   MV_MV22_CV1 : PlantItem := (CW := 2#0000_0000_0000_0000_0000_0000_1000_0001, DriveBits := 1);   // MV22_CV1
   MV_MV22_CV1_RawOutput : ALIAS FOR Remote_IO:12:O.Data.11;   // MV_MV22_CV1 MV22 coolant SOV
   MV_MV22_Filling_Pulse : BOOL;
   MV_MV22_Filling_PulseLevel : DINT := 252;
   MV_MV22_LTX07_AI : PlantItem := (CW := 2#0000_0000_0000_0000_1000_0000_0000_0000, CheckTime := 10, CheckTimer := 10, Scaled := 5.5534997, RawInput := 7064.0);   // MV22_LTX07
   MV_MV22_LTX07_AI_RawInput : ALIAS FOR Remote_IO:10:I.Ch05Data;   // Real Analog Input , Do Not Use In Code
   MV_MV22_LTX07_TrueLevel : REAL := 251.42085;
   MV_MV22_LTX07_TruePressure : REAL := 5.5534997;
   MV_MV22_Open_Vent_ALRM : ALARM_DIGITAL;
   MV_MV22_ProxiesOK : BOOL;
   MV_MV22_PTX01_AI : PlantItem := (CW := 2#0000_0000_0000_0000_1000_0000_0000_0000, CheckTime := 10, CheckTimer := 10, Scaled := -0.060749996, RawInput := 3946.0);   // MV22_PTX01
   MV_MV22_PTX01_AI_RawInput : ALIAS FOR Remote_IO:10:I.Ch02Data;   // Real Analog Input , Do Not Use In Code
   MV_MV22_PurgeAfterCIP : BOOL;
   MV_MV22_RTD1_AI : PlantItem := (CW := 2#0000_0000_0000_0000_1000_0000_0000_0000, CheckTime := 10, CheckTimer := 10, Scaled := -0.19999886, RawInput := -2.0);   // MV22_RTD1
   MV_MV22_RTD1_AI_RawInput : ALIAS FOR Remote_IO:5:I.Ch3Data;   // Real Analog Input , Do Not Use In Code
   MV_MV22_TP_CaskDepressure : BOOL;
   MV_MV22_TP_CaskEmptying : BOOL;
   MV_MV22_TP_CaskFilling : BOOL;
   MV_MV22_TP_CaskPreEmptyPressure : BOOL;
   MV_MV22_TP_CaskPrePressure : BOOL;
   MV_MV22_TP_CaskPressureDelay : BOOL;
   MV_MV22_TP_CaskPurgeFromTop : BOOL;
   MV_MV22_TP_CaskReadyToFill : BOOL;
   MV_MV22_TP_CaskStorage : BOOL;
   MV_MV22_TP_CO2_Debounce_Timer : TIMER := (PRE := 5000);
   MV_MV22_TP_CO2_Debounce_Timer_1 : TIMER := (PRE := 5000);
   MV_MV22_TP_CO2_HSL_Pressure : REAL := 16.0;
   MV_MV22_TP_CO2_HSL_Storage : REAL := 10.5;
   MV_MV22_TP_CO2_HSL_Timer : TIMER := (PRE := 5000, ACC := 5000, EN := 1, DN := 1);
   MV_MV22_TP_CO2_LSL_pressure : DINT := 9;
   MV_MV22_TP_CO2_LSL_pressure_1 : REAL := 2.0;
   MV_MV22_TP_CO2_LSL_storage : REAL := 9.5;
   MV_MV22_TP_CO2_LSL_Timer : TIMER := (PRE := 5000);
   MV_MV22_TP_CO2_Overshoot_pressure : DINT := 4;
   MV_MV22_TP_CO2_Pulse_Debounce_Timer : TIMER := (PRE := 5000);
   MV_MV22_TP_Command : DINT;
   MV_MV22_TP_DAL_Chase_Cask : BOOL;
   MV_MV22_TP_DAL_Chase_KB : BOOL;
   MV_MV22_TP_DAL_Chase_Time : TIMER := (PRE := 90000);
   MV_MV22_TP_Dirty : BOOL;
   MV_MV22_TP_DrainDown : BOOL;
   MV_MV22_TP_Emptying_Level_Setpoint : REAL := -260.0;
   MV_MV22_TP_Error_String : STRING;
   MV_MV22_TP_Faulted : BOOL;
   MV_MV22_TP_Fill_Pulse_OFF_Timer : TIMER := (PRE := 15000);
   MV_MV22_TP_Fill_Pulse_ON_Timer : TIMER := (PRE := 30000);
   MV_MV22_TP_Held : BOOL;
   MV_MV22_TP_Idle : BOOL;
   MV_MV22_TP_Initial_DAL_Chase_Cask : BOOL;
   MV_MV22_TP_Initial_DAL_Chase_KB : BOOL;
   MV_MV22_TP_KBDepressure : BOOL;
   MV_MV22_TP_KBEmptying : BOOL;
   MV_MV22_TP_KBFilling : BOOL;
   MV_MV22_TP_KBFilling_M : BOOL;
   MV_MV22_TP_KBFillingBuildPressure : BOOL;
   MV_MV22_TP_KBPreEmptyPressure : BOOL;
   MV_MV22_TP_KBPrePressurise : BOOL;
   MV_MV22_TP_KBPurgeFromTop : BOOL;
   MV_MV22_TP_KBPurgeTimer : TIMER;
   MV_MV22_TP_KBStorage : BOOL := 1;
   MV_MV22_TP_LowerLimit : REAL := 8.0;
   MV_MV22_TP_NotIdle : BOOL := 1;
   MV_MV22_TP_ONS : BOOL;
   MV_MV22_TP_ONS_1 : BOOL;
   MV_MV22_TP_PrePressure : BOOL;
   MV_MV22_TP_Prompt : DINT := 2;
   MV_MV22_TP_Proxy_Delay_Made : TIMER := (PRE := 2000);
   MV_MV22_TP_Proxy_Delay_NOT_MADE : TIMER := (PRE := 2000, ACC := 2000, EN := 1, DN := 1);
   MV_MV22_TP_Pulse : BOOL;
   MV_MV22_TP_ReadyToFillKB : BOOL;
   MV_MV22_TP_ReadyToFillKB_M : BOOL;
   MV_MV22_TP_Running : BOOL := 1;
   MV_MV22_TP_SeatClean_Delay : TIMER;
   MV_MV22_TP_SeatClean_Pulse : TIMER;
   MV_MV22_TP_Setpoint : REAL := 10.0;
   MV_MV22_TP_Status : DINT := 1;   // 0 = Idle, 1 = Running, 2 = Held, 3 = Faulted
   MV_MV22_TP_Step : DINT := 50;
   MV_MV22_TP_Steptime : DINT := 3562924;
   MV_MV22_TP_Steptime_String : STRING := '989:42:06';
   MV_MV22_TP_Steptime_String_1 : STRING;
   MV_MV22_TP_SteptimeRunning : DINT := 11;
   MV_MV22_TP_TimeLeft : DINT;
   MV_MV22_TP_TimeLeft_msec : DINT := 1;
   MV_MV22_TP_TimeLeftStr : STRING;
   MV_MV22_TP_UpperLimit : REAL := 12.0;
   MV_MV22_TP_Vent : BOOL;
   MV_MV22_TP_VentPressure : REAL;
   MV_MV22_TPLastStep : DINT := 50;
   MV_MV22_Transfer_StartLevel : REAL;
   MV_MV22_Transferred_Level : REAL := 95.31006;
   MV_MV22R : PlantItem := (CW := 2#0000_0000_0000_0010_0000_1100_0100_0001, CheckTime := 8, DriveBits := 1);   // MV22R
   MV_MV22R_ALARM : ALARM_DIGITAL;
   MV_MV22R_D : ALIAS FOR Remote_IO:14:O.Data.11;   // Rouser drive MV22
   MV_MV22R_R : ALIAS FOR Remote_IO:15:I.Data.27;   // MV22 Rouser running signal
   MV_MV23_CV1 : PlantItem;   // MV23_CV1
   MV_MV23_CV1_RawOutput : ALIAS FOR Remote_IO:12:O.Data.12;   // MV_MV23_CV1 MV23 coolant SOV
   MV_MV23_RTD1_AI : PlantItem := (CW := 2#0000_0000_0000_0000_1000_0000_0000_0000, CheckTime := 10, CheckTimer := 10, Scaled := 8.300001, RawInput := 83.0);   // MV23_RTD1
   MV_MV23_RTD1_AI_RawInput : ALIAS FOR Remote_IO:5:I.Ch4Data;   // Real Analog Input , Do Not Use In Code
   MV_MV23R : PlantItem := (CW := 2#0000_0000_0000_0010_0000_1100_0000_0000, CheckTime := 8, CheckTimer := 8);   // MV23R
   MV_MV23R_ALARM : ALARM_DIGITAL;
   MV_MV23R_D : ALIAS FOR Remote_IO:14:O.Data.12;   // Rouser drive MV23
   MV_MV23R_R : ALIAS FOR Remote_IO:15:I.Data.28;   // MV23 Rouser running signal
   MV_MV2_CV1 : PlantItem;   // MV2_CV1
   MV_MV2_CV1_RawOutput : ALIAS FOR Remote_IO:11:O.Data.1;   // MV_MV2_CV1
   MV_MV2_RTD1_AI : PlantItem := (CW := 2#0000_0000_0000_0000_1000_0000_0000_0000, CheckTime := 10, CheckTimer := 10, Scaled := 8.200001, RawInput := 82.0);   // MV2_RTD1
   MV_MV2_RTD1_AI_RawInput : ALIAS FOR Remote_IO:1:I.Ch1Data;   // Real Analog Input , Do Not Use In Code
   MV_MV2R : PlantItem := (CW := 2#0000_0000_0000_0011_0000_1100_0000_0000, CheckTime := 8, CheckTimer := 8);   // MV2R
   MV_MV2R_ALARM : ALARM_DIGITAL;
   MV_MV2R_ALM : ALARM_DIGITAL;
   MV_MV2R_D : ALIAS FOR Remote_IO:13:O.Data.1;
   MV_MV2R_R : ALIAS FOR Remote_IO:15:I.Data.1;   // MV2 Rouser running signal
   MV_MV30_CV1 : PlantItem;   // MV30_CV1
   MV_MV30_CV1_RawOutput : ALIAS FOR Remote_IO:12:O.Data.3;   // MV_MV30_CV1 MV30 coolant SOV
   MV_MV30_RTD1_AI : PlantItem := (CW := 2#0000_0000_0000_0000_1000_0000_0000_0000, CheckTime := 10, CheckTimer := 10, Scaled := 21.900002, RawInput := 219.0);   // MV30_RTD1
   MV_MV30_RTD1_AI_RawInput : ALIAS FOR Remote_IO:4:I.Ch1Data;   // Real Analog Input , Do Not Use In Code
   MV_MV30R : PlantItem := (CW := 2#0000_0000_0000_0010_0000_1100_0000_0000, CheckTime := 8, CheckTimer := 8);   // MV30R
   MV_MV30R_ALARM : ALARM_DIGITAL;
   MV_MV30R_D : ALIAS FOR Remote_IO:14:O.Data.3;   // Rouser drive MV30
   MV_MV30R_R : ALIAS FOR Remote_IO:15:I.Data.19;   // MV30 Rouser running signal
   MV_MV31_CV1 : PlantItem;   // MV31_CV1
   MV_MV31_CV1_RawOutput : ALIAS FOR Remote_IO:12:O.Data.4;   // MV_MV31_CV1 MV31coolant SOV
   MV_MV31_RTD1_AI : PlantItem := (CW := 2#0000_0000_0000_0000_1000_0000_0000_0000, CheckTime := 10, CheckTimer := 10, Scaled := 6.300001, RawInput := 63.0);   // MV31_RTD1
   MV_MV31_RTD1_AI_RawInput : ALIAS FOR Remote_IO:4:I.Ch2Data;   // Real Analog Input , Do Not Use In Code
   MV_MV31R : PlantItem := (CW := 2#0000_0000_0000_0010_0000_1100_0000_0000, CheckTime := 8, CheckTimer := 8);   // MV31R
   MV_MV31R_ALARM : ALARM_DIGITAL;
   MV_MV31R_D : ALIAS FOR Remote_IO:14:O.Data.4;   // Rouser drive MV31
   MV_MV31R_R : ALIAS FOR Remote_IO:15:I.Data.20;   // MV31 Rouser running signal
   MV_MV32_CV1 : PlantItem;   // MV32_CV1
   MV_MV32_CV1_RawOutput : ALIAS FOR Remote_IO:12:O.Data.5;   // MV_MV32_CV1 MV32 coolant SOV
   MV_MV32_RTD1_AI : PlantItem := (CW := 2#0000_0000_0000_0000_1000_0000_0000_0000, CheckTime := 10, CheckTimer := 10, Scaled := 22.0, RawInput := 220.0);   // MV32_RTD1
   MV_MV32_RTD1_AI_RawInput : ALIAS FOR Remote_IO:4:I.Ch3Data;   // Real Analog Input , Do Not Use In Code
   MV_MV32R : PlantItem := (CW := 2#0000_0000_0000_0010_0000_1100_0000_0000, CheckTime := 8, CheckTimer := 8);   // MV32R
   MV_MV32R_ALARM : ALARM_DIGITAL;
   MV_MV32R_D : ALIAS FOR Remote_IO:14:O.Data.5;   // Rouser drive MV32
   MV_MV32R_R : ALIAS FOR Remote_IO:15:I.Data.21;   // MV32 Rouser running signal
   MV_MV33_CV1 : PlantItem;   // MV33_CV1
   MV_MV33_CV1_RawOutput : ALIAS FOR Remote_IO:12:O.Data.6;   // MV_MV33_CV1 MV33 coolant SOV
   MV_MV33_RTD1_AI : PlantItem := (CW := 2#0000_0000_0000_0000_1000_0000_0000_0000, CheckTime := 10, CheckTimer := 10, Scaled := 8.1, RawInput := 81.0);   // MV33_RTD1
   MV_MV33_RTD1_AI_RawInput : ALIAS FOR Remote_IO:4:I.Ch4Data;   // Real Analog Input , Do Not Use In Code
   MV_MV33R : PlantItem := (CW := 2#0000_0000_0000_0010_0000_1100_0000_0000, CheckTime := 8, CheckTimer := 8);   // MV33R
   MV_MV33R_ALARM : ALARM_DIGITAL;
   MV_MV33R_D : ALIAS FOR Remote_IO:14:O.Data.6;   // Rouser drive MV33
   MV_MV33R_R : ALIAS FOR Remote_IO:15:I.Data.22;   // MV33 Rouser running signal
   MV_MV34_CV1 : PlantItem;   // MV34_CV1
   MV_MV34_CV1_RawOutput : ALIAS FOR Remote_IO:12:O.Data.7;   // MV_MV34_CV1 MV34 coolant SOV
   MV_MV34_RTD1_AI : PlantItem := (CW := 2#0000_0000_0000_0000_1000_0000_0000_0000, CheckTime := 10, CheckTimer := 10, Scaled := 22.100002, RawInput := 221.0);   // MV34_RTD1
   MV_MV34_RTD1_AI_RawInput : ALIAS FOR Remote_IO:4:I.Ch5Data;   // Real Analog Input , Do Not Use In Code
   MV_MV34R : PlantItem := (CW := 2#0000_0000_0000_0010_0000_1100_0000_0000, CheckTime := 8, CheckTimer := 8);   // MV34R
   MV_MV34R_ALARM : ALARM_DIGITAL;
   MV_MV34R_D : ALIAS FOR Remote_IO:14:O.Data.7;   // Rouser drive MV34
   MV_MV34R_R : ALIAS FOR Remote_IO:15:I.Data.23;   // MV34 Rouser running signal
   MV_MV35_CV1 : PlantItem;   // MV35_CV1
   MV_MV35_CV1_RawOutput : ALIAS FOR Remote_IO:12:O.Data.8;   // MV_MV35_CV1 MV35 coolant SOV
   MV_MV35_RTD1_AI : PlantItem := (CW := 2#0000_0000_0000_0000_1000_0000_0000_0000, CheckTime := 10, CheckTimer := 10, Scaled := 22.8, RawInput := 228.0);   // MV35_RTD1
   MV_MV35_RTD1_AI_RawInput : ALIAS FOR Remote_IO:5:I.Ch0Data;   // Real Analog Input , Do Not Use In Code
   MV_MV35R : PlantItem := (CW := 2#0000_0000_0000_0010_0000_1100_0000_0000, CheckTime := 8, CheckTimer := 8);   // MV35R
   MV_MV35R_ALARM : ALARM_DIGITAL;
   MV_MV35R_D : ALIAS FOR Remote_IO:14:O.Data.8;   // Rouser drive MV35
   MV_MV35R_R : ALIAS FOR Remote_IO:15:I.Data.24;   // MV35 Rouser running signal
   MV_MV36_AV01 : PlantItem;   // MV36_AV01
   MV_MV36_AV01_RawOutput : ALIAS FOR Remote_IO:16:O.Data.0;   // MV_MV36_AV01
   MV_MV36_TTX01_AI : PlantItem := (CW := 2#0000_0000_0000_0000_1000_0000_0000_0000, CheckTime := 10, CheckTimer := 10, Scaled := 8.096876, RawInput := 9791.0);   // MV36_TTX01
   MV_MV36_TTX01_AI_RawInput : ALIAS FOR Remote_IO:7:I.Ch00Data;   // Real Analog Input , Do Not Use In Code
   MV_MV37_AV01 : PlantItem := (CW := 2#0000_0000_0000_0000_0000_0000_0010_0000);   // MV37_AV01
   MV_MV37_AV01_RawOutput : ALIAS FOR Remote_IO:16:O.Data.1;   // MV_MV37_AV01 MV37 coolant SOV
   MV_MV37_TTX01_AI : PlantItem := (CW := 2#0000_0000_0000_0000_1000_0000_0000_0000, CheckTime := 10, CheckTimer := 10, Scaled := -1.4093752, RawInput := 6749.0);   // MV37_TTX01
   MV_MV37_TTX01_AI_RawInput : ALIAS FOR Remote_IO:7:I.Ch01Data;   // Real Analog Input , Do Not Use In Code
   MV_MV38_AV01 : PlantItem;   // MV38_AV01
   MV_MV38_AV01_RawOutput : ALIAS FOR Remote_IO:16:O.Data.2;   // MV_MV38_AV01 MV38 coolant SOV
   MV_MV38_TTX01_AI : PlantItem := (CW := 2#0000_0000_0000_0000_1000_0000_0000_0000, CheckTime := 10, CheckTimer := 10, Scaled := 8.1, RawInput := 9792.0);   // MV38_TTX01
   MV_MV38_TTX01_AI_RawInput : ALIAS FOR Remote_IO:7:I.Ch02Data;   // Real Analog Input , Do Not Use In Code
   MV_MV39_AV01 : PlantItem;   // MV39_AV01
   MV_MV39_AV01_RawOutput : ALIAS FOR Remote_IO:16:O.Data.3;   // MV_MV39_AV01 MV39 coolant SOV
   MV_MV39_TTX01_AI : PlantItem := (CW := 2#0000_0000_0000_0000_1000_0000_0000_0000, CheckTime := 10, CheckTimer := 10, Scaled := -1.4437494, RawInput := 6738.0);   // MV39_TTX01
   MV_MV39_TTX01_AI_RawInput : ALIAS FOR Remote_IO:7:I.Ch03Data;   // Real Analog Input , Do Not Use In Code
   MV_MV3_CV1 : PlantItem;   // MV3_CV1
   MV_MV3_CV1_RawOutput : ALIAS FOR Remote_IO:11:O.Data.2;   // MV_MV3_CV1 MV3 coolant SOV
   MV_MV3_RTD1_AI : PlantItem := (CW := 2#0000_0000_0000_0000_1000_0000_0000_0000, CheckTime := 10, CheckTimer := 10, Scaled := 8.1, RawInput := 81.0);   // MV3_RTD1
   MV_MV3_RTD1_AI_RawInput : ALIAS FOR Remote_IO:1:I.Ch2Data;   // Real Analog Input , Do Not Use In Code
   MV_MV3R : PlantItem := (CW := 2#0000_0000_0000_0010_0000_1100_0000_0000, CheckTime := 8, CheckTimer := 8);   // MV3R
   MV_MV3R_ALARM : ALARM_DIGITAL;
   MV_MV3R_D : ALIAS FOR Remote_IO:13:O.Data.2;   // Rouser drive MV3
   MV_MV3R_R : ALIAS FOR Remote_IO:15:I.Data.2;   // MV3 Rouser running signal
   MV_MV40_AV01 : PlantItem;   // MV40_AV01
   MV_MV40_AV01_RawOutput : ALIAS FOR Remote_IO:16:O.Data.4;   // MV_MV40_AV01 MV40 coolant SOV
   MV_MV40_TTX01_AI : PlantItem := (CW := 2#0000_0000_0000_0000_1000_0000_0000_0000, CheckTime := 10, CheckTimer := 10, Scaled := 7.7562504, RawInput := 9682.0);   // MV40_TTX01
   MV_MV40_TTX01_AI_RawInput : ALIAS FOR Remote_IO:7:I.Ch04Data;   // Real Analog Input , Do Not Use In Code
   MV_MV41_AV01 : PlantItem;   // MV41_AV01
   MV_MV41_AV01_RawOutput : ALIAS FOR Remote_IO:16:O.Data.5;   // MV_MV41_AV01 MV41 coolant SOV
   MV_MV41_TTX01_AI : PlantItem := (CW := 2#0000_0000_0000_0000_1000_0000_0000_0000, CheckTime := 10, CheckTimer := 10, Scaled := 7.846876, RawInput := 9711.0);   // MV41_TTX01
   MV_MV41_TTX01_AI_RawInput : ALIAS FOR Remote_IO:7:I.Ch05Data;   // Real Analog Input , Do Not Use In Code
   MV_MV42_AV01 : PlantItem;   // MV42_AV01
   MV_MV42_AV01_RawOutput : ALIAS FOR Remote_IO:16:O.Data.6;   // MV_MV42_AV01 MV42 coolant SOV
   MV_MV42_TTX01_AI : PlantItem := (CW := 2#0000_0000_0000_0000_1000_0000_0000_0000, CheckTime := 10, CheckTimer := 10, Scaled := 21.015625, RawInput := 13925.0);   // MV42_TTX01
   MV_MV42_TTX01_AI_RawInput : ALIAS FOR Remote_IO:7:I.Ch06Data;   // Real Analog Input , Do Not Use In Code
   MV_MV43_AV01 : PlantItem;   // MV43_AV01
   MV_MV43_AV01_RawOutput : ALIAS FOR Remote_IO:16:O.Data.7;   // MV_MV43_AV01 MV43 coolant SOV
   MV_MV43_TTX01_AI : PlantItem := (CW := 2#0000_0000_0000_0000_1000_0000_0000_0000, CheckTime := 10, CheckTimer := 10, Scaled := 21.221876, RawInput := 13991.0);   // MV43_TTX01
   MV_MV43_TTX01_AI_RawInput : ALIAS FOR Remote_IO:7:I.Ch07Data;   // Real Analog Input , Do Not Use In Code
   MV_MV44_AV01 : PlantItem;   // MV44_AV01
   MV_MV44_AV01_RawOutput : ALIAS FOR Remote_IO:16:O.Data.8;   // MV_MV44_AV01 MV44 coolant SOV
   MV_MV44_TTX01_AI : PlantItem := (CW := 2#0000_0000_0000_0000_1000_0000_0000_0000, CheckTime := 10, CheckTimer := 10, Scaled := 21.075, RawInput := 13944.0);   // MV44_TTX01
   MV_MV44_TTX01_AI_RawInput : ALIAS FOR Remote_IO:7:I.Ch08Data;   // Real Analog Input , Do Not Use In Code
   MV_MV45_AV01 : PlantItem;   // MV45_AV01
   MV_MV45_AV01_RawOutput : ALIAS FOR Remote_IO:16:O.Data.9;   // MV_MV45_AV01 MV45 coolant SOV
   MV_MV45_TTX01_AI : PlantItem := (CW := 2#0000_0000_0000_0000_1000_0000_0000_0000, CheckTime := 10, CheckTimer := 10, Scaled := 7.778126, RawInput := 9689.0);   // MV45_TTX01
   MV_MV45_TTX01_AI_RawInput : ALIAS FOR Remote_IO:7:I.Ch09Data;   // Real Analog Input , Do Not Use In Code
   MV_MV46_AV01 : PlantItem;   // MV46_AV01
   MV_MV46_AV01_RawOutput : ALIAS FOR Remote_IO:16:O.Data.10;   // MV_MV46_AV01 MV46 coolant SOV
   MV_MV46_TTX01_AI : PlantItem := (CW := 2#0000_0000_0000_0000_1000_0000_0000_0000, CheckTime := 10, CheckTimer := 10, Scaled := 21.25625, RawInput := 14002.0);   // MV46_TTX01
   MV_MV46_TTX01_AI_RawInput : ALIAS FOR Remote_IO:7:I.Ch10Data;   // Real Analog Input , Do Not Use In Code
   MV_MV47_AV01 : PlantItem := (CW := 2#0000_0000_0000_0000_0000_0000_1000_0001, DriveBits := 1);   // MV47_AV01
   MV_MV47_AV01_RawOutput : ALIAS FOR Remote_IO:16:O.Data.11;   // MV_MV47_AV01 MV47 coolant SOV
   MV_MV47_TTX01_AI : PlantItem := (CW := 2#0000_0000_0000_0000_1000_0000_0000_0000, CheckTime := 10, CheckTimer := 10, Scaled := -1.2468748, RawInput := 6801.0);   // MV47_TTX01
   MV_MV47_TTX01_AI_RawInput : ALIAS FOR Remote_IO:7:I.Ch11Data;   // Real Analog Input , Do Not Use In Code
   MV_MV4_CV1 : PlantItem;   // MV4_CV1
   MV_MV4_CV1_RawOutput : ALIAS FOR Remote_IO:11:O.Data.3;   // MV_MV4_CV1 MV4 coolant SOV
   MV_MV4_RTD1_AI : PlantItem := (CW := 2#0000_0000_0000_0000_1000_0000_0000_0000, CheckTime := 10, CheckTimer := 10, Scaled := 8.0, RawInput := 80.0);   // MV4_RTD1
   MV_MV4_RTD1_AI_RawInput : ALIAS FOR Remote_IO:1:I.Ch3Data;   // Real Analog Input , Do Not Use In Code
   MV_MV4R : PlantItem := (CW := 2#0000_0000_0000_0010_0000_1100_0000_0000, CheckTime := 8, CheckTimer := 8);   // MV4R
   MV_MV4R_ALARM : ALARM_DIGITAL;
   MV_MV4R_D : ALIAS FOR Remote_IO:13:O.Data.3;   // Rouser drive MV4
   MV_MV4R_R : ALIAS FOR Remote_IO:15:I.Data.3;   // MV4 Rouser running signal
   MV_MV5_CV1 : PlantItem;   // MV5_CV1
   MV_MV5_CV1_RawOutput : ALIAS FOR Remote_IO:11:O.Data.4;   // MV_MV5_CV1 MV5 coolant SOV
   MV_MV5_RTD1_AI : PlantItem := (CW := 2#0000_0000_0000_0000_1000_0000_0000_0000, CheckTime := 10, CheckTimer := 10, Scaled := 8.200001, RawInput := 82.0);   // MV5_RTD1
   MV_MV5_RTD1_AI_RawInput : ALIAS FOR Remote_IO:1:I.Ch4Data;   // Real Analog Input , Do Not Use In Code
   MV_MV5R : PlantItem := (CW := 2#0000_0000_0000_0010_0000_1100_0000_0000, CheckTime := 8, CheckTimer := 8);   // MV5R
   MV_MV5R_ALARM : ALARM_DIGITAL;
   MV_MV5R_D : ALIAS FOR Remote_IO:13:O.Data.4;   // Rouser drive MV5
   MV_MV5R_R : ALIAS FOR Remote_IO:15:I.Data.4;   // MV5 Rouser running signal
   MV_MV6_CV1 : PlantItem;   // MV6_CV1
   MV_MV6_CV1_RawOutput : ALIAS FOR Remote_IO:11:O.Data.5;   // MV_MV6_CV1 MV6 coolant SOV
   MV_MV6_RTD1_AI : PlantItem := (CW := 2#0000_0000_0000_0000_1000_0000_0000_0000, CheckTime := 10, CheckTimer := 10, Scaled := 25.100002, RawInput := 251.0);   // MV6_RTD1
   MV_MV6_RTD1_AI_RawInput : ALIAS FOR Remote_IO:1:I.Ch5Data;   // Real Analog Input , Do Not Use In Code
   MV_MV6R : PlantItem := (CW := 2#0000_0000_0000_0010_0000_1100_0000_0000, CheckTime := 8, CheckTimer := 8);   // MV6R
   MV_MV6R_ALARM : ALARM_DIGITAL;
   MV_MV6R_D : ALIAS FOR Remote_IO:13:O.Data.5;   // Rouser drive MV6
   MV_MV6R_R : ALIAS FOR Remote_IO:15:I.Data.5;   // MV6 Rouser running signal
   MV_MV7_CV1 : PlantItem;   // MV7_CV1
   MV_MV7_CV1_RawOutput : ALIAS FOR Remote_IO:11:O.Data.6;   // MV_MV7_CV1 MV7 coolant SOV
   MV_MV7_RTD1_AI : PlantItem := (CW := 2#0000_0000_0000_0000_1000_0000_0000_0000, CheckTime := 10, CheckTimer := 10, Scaled := 8.200001, RawInput := 82.0);   // MV7_RTD1
   MV_MV7_RTD1_AI_RawInput : ALIAS FOR Remote_IO:2:I.Ch0Data;   // Real Analog Input , Do Not Use In Code
   MV_MV7R : PlantItem := (CW := 2#0000_0000_0000_0010_0000_1100_0000_0000, CheckTime := 8, CheckTimer := 8);   // MV7R
   MV_MV7R_ALARM : ALARM_DIGITAL;
   MV_MV7R_D : ALIAS FOR Remote_IO:13:O.Data.6;   // Rouser drive MV7
   MV_MV7R_R : ALIAS FOR Remote_IO:15:I.Data.6;   // MV7 Rouser running signal
   MV_MV8_CV1 : PlantItem := (CW := 2#0000_0000_0000_0000_0000_0000_1000_0001, DriveBits := 1);   // MV8_CV1
   MV_MV8_CV1_RawOutput : ALIAS FOR Remote_IO:11:O.Data.7;   // MV_MV8_CV1 MV8 coolant SOV
   MV_MV8_RTD1_AI : PlantItem := (CW := 2#0000_0000_0000_0000_1000_0000_0000_0000, CheckTime := 10, CheckTimer := 10, Scaled := 9.700001, RawInput := 97.0);   // MV8_RTD1
   MV_MV8_RTD1_AI_RawInput : ALIAS FOR Remote_IO:2:I.Ch1Data;   // Real Analog Input , Do Not Use In Code
   MV_MV8R : PlantItem := (CW := 2#0000_0000_0000_0010_0000_1100_0000_0000, CheckTime := 8, CheckTimer := 8);   // MV8R
   MV_MV8R_ALARM : ALARM_DIGITAL;
   MV_MV8R_D : ALIAS FOR Remote_IO:13:O.Data.7;   // Rouser drive MV8
   MV_MV8R_R : ALIAS FOR Remote_IO:15:I.Data.7;   // MV8 Rouser running signal
   MV_MV9_CV1 : PlantItem := (CW := 2#0000_0000_0000_0000_0000_0000_0010_0000);   // MV9_CV1
   MV_MV9_CV1_RawOutput : ALIAS FOR Remote_IO:11:O.Data.8;   // MV_MV9_CV1 MV9 coolant SOV
   MV_MV9_RTD1_AI : PlantItem := (CW := 2#0000_0000_0000_0000_1000_0000_0000_0000, CheckTime := 10, CheckTimer := 10, Scaled := 26.400002, RawInput := 264.0);   // MV9_RTD1
   MV_MV9_RTD1_AI_RawInput : ALIAS FOR Remote_IO:2:I.Ch2Data;   // Real Analog Input , Do Not Use In Code
   MV_MV9R : PlantItem := (CW := 2#0000_0000_0000_0010_0000_1100_0000_0000, CheckTime := 8, CheckTimer := 8);   // MV9R
   MV_MV9R_ALARM : ALARM_DIGITAL;
   MV_MV9R_D : ALIAS FOR Remote_IO:13:O.Data.8;   // Rouser drive MV9
   MV_MV9R_R : ALIAS FOR Remote_IO:15:I.Data.8;   // MV9 Rouser running signal
   MV_N101 : INT[255] := ([0] := 152, [1] := -15, [2] := -15, [3] := 1680, [4] := 5280, [5] := 2950, [6] := 463, [7] := 124, [8] := 7, [9] := 3, [10] := 110, [11] := -13);   // AT INT Fermentation control integer workspace
        [1]   // Setpoint at previous breakpoint
        [4]   // Next breakpoint time
        [6]   // Temporary result register
        [5]   // Time since last B.P in 1/10 hour
        [3]   // Previous breakpoint time
        [0]   // Attemporation Control Loop Current Vessel File Pointer
        [7]   // Pointer to vessel's data file
        [8]   // Number of open cooling valves
        [11]   // Temp.register
        [2]   // Setpoint at next breakpoint
        [9]   // Rouser operation temperature
   MV_N104 : INT[255] := ([0] := -32768, [1] := -32768, [2] := -32768, [3] := -32768, [4] := -32768, [5] := -32768, [6] := -32768, [7] := -32768, [8] := -32768, [9] := -32768, [10] := -32768, [11] := -32768, [12] := -32768, [13] := -32768, [14] := -32768, [15] := -32768, [16] := -32768, [17] := -32768, [18] := -32768, [19] := -32768, [20] := -32768, [21] := -32768, [22] := -32768, [23] := -32768, [24] := -32768);   // MV_PC_BUF PC>PLC Attemporation Control Command Buf fer File
        [10]   // PC>PLC FV System Command Buffer Breakpoint E Temperature Setpoint
        [12]   // PC>PLC FV System Command Buffer Breakpoint F Temperature Setpoint
        [14]   // PC>PLC FV System Command Buffer Breakpoint G Temperature Setpoint
        [1]   // PC>PLC Attemporation System Command Buffer Breakpoint A Time
        [15]   // PC>PLC FV System Command Buffer Profile Control / Configuration Flags
        [15].6   // FV System PC Command Buffer Control Flags 1=Wait for yeast required
        [2]   // PC>PLC FV System Command Buffer Breakpoint A Temperature Setpoint
        [4]   // PC>PLC FV System Command Buffer Breakpoint B Temperature Setpoint
        [6]   // PC>PLC FV System Command Buffer Breakpoint C Temperature Setpoint
        [15].4   // FV System PC Command Buffer Control Flags 1=Ageing Profile
        [8]   // PC>PLC FV System Command Buffer Breakpoint D Temperature Setpoint
        [23]   // PC>PLC AT System Command Buffer Command Type 1=Start,2=Stop 3=Modify Control
        [0]   // PC>PLC Attempotation System Vessel Number 29-56,94 = MV1-MV23 336-347 = MV36-47
        [15].5   // FV System PC Command Buffer Control Flags 1=Conditioning Profile
        [11]   // PC>PLC FV System Command Buffer Breakpoint F Time
        [13]   // PC>PLC FV System Command Buffer Breakpoint G Time
        [24]   // Attemporation System PC Command Buffer Phase Number
        [16]   // PC>PLC FV System Command Buffer PC Private Flags
        [3]   // PC>PLC FV System Command Buffer Breakpoint B Time
        [5]   // PC>PLC FV System Command Buffer Breakpoint C Time
        [7]   // PC>PLC FV System Command Buffer Breakpoint D Time
        [9]   // PC>PLC FV System Command Buffer Breakpoint E Time
   MV_N105 : INT[255] := ([0] := 1025, [1] := 116, [3] := 45, [4] := 114);   // ROUSE_CTRL Rouser control progr am working regs
        [2]   // PC>PLC Rouser control Vessel number to be set to timed mode
        [0].0   // Rouser control 1 minute latch
        [0].10   // Rouser Control Hourly Latch
        [0].2   // Rouser Control Daily latch synchroniser
        [0].9   // Rouser Control Hourly latch synchroniser
        [4]   // Rouse control PC timed rouse request vessel pointer
        [1]   // Rouser control current vessel data file pointer
        [0].3   // Rouser Control Daily Latch
        [3]   // PC>PLC Rouser control Timed rouse duration
        [0].4   // Rouser control 1 minute latch synchroniser
   MV_N105_0_1_Output_Bit : BOOL;
   MV_N105_0_6_Output_Bit : BOOL;
   MV_N105_0_7_Output_Bit : BOOL;
   MV_N105_0_8_Output_Bit : BOOL;
   MV_N106 : INT[255] := ([0] := 33, [2] := 80, [3] := 1680, [4] := 80, [5] := 3360, [6] := 80, [7] := 5040, [8] := 80, [9] := 6720, [10] := 80, [11] := 8400, [12] := 80, [13] := 32767, [14] := 80, [15] := 148, [17] := -32767, [18] := -32767, [19] := 1680, [20] := 3171, [22] := 4639, [23] := 1, [24] := 10, [25] := 82, [26] := 80, [27] := 3171, [29] := 2, [30] := 24, [32] := 2, [34] := 2, [42] := 25640);   // ROUSE_BUFF Rouser control vesse l data buffer
        [24]   // Phase 0=off 8=Wait yeast 10=Maturation 11to16=Conditioning
        [32]   // Rouser control mode 0=Off 1=Continuous 2=Daily 3=Timed 4=Hourly
        [30].2   // Rouse required due to high temperature
        [29].1   // Current vessel deferred chilling enabled flag
        [30].0   // Current vessel cooling valve required to open
        [34]   // Saved rouser mode of operation
        [27]   // Current vessel elapsed time
        [15].7   // Profile control flag Rousing enabled
        [25]   // ACTUAL TEMPERATURE -DEGREES 'C'*10
        [30].1   // Rouser to run
        [31]   // Rouser run time remaining (minutes)
   MV_N110 : INT[255] := ([0] := 347, [2] := 100, [3] := 1200, [4] := 100, [5] := 1680, [6] := -15, [7] := 5280, [8] := -15, [9] := 7210, [10] := -15, [11] := 8340, [12] := -15, [13] := 32767, [14] := -15, [15] := 164, [17] := -32767, [18] := -32767, [19] := 1680, [20] := 1200, [21] := 2981, [22] := 6282, [23] := 1, [24] := 13, [25] := -13, [26] := -15, [27] := 4630, [29] := 257, [30] := 123, [32] := 2, [34] := 2, [40] := 2);   // MV DATA 0 CURRENT FV DATA
        [15].5   // Profile Control Flags : This is a Conditioning Profile
        [24]   // Phase 0=off 8=Wait yeast 9=Wait Fill 10=Maturation 11to16=Conditioning
        [15].9   // Current vessel deferred chilling manual override
        [22]   // Current FV total residence time
        [29].0   // PC TO SAVE TEMPERATURE DATA
        [40]   // Vessel RoutingStatus 0=Clean,1=Filling,2= Beer,3=Packng1,4=Pac kng2,5=Packng3,6=Ven ting,7=Dirty,8=CIP
        [15].4   // Profile Control Flags : This is a Maturation Profile
        [1]   // TEMPERATURE BREAKPOINT A. TIME 1/10 HOURS(ALWAYS=0)
        [11]   // TEMPERATURE BREAKPOINT F. TIME 1/10 HOURS(ALWAYS=0)
        [29].1   // Current vessel deferred chilling enabled flag
        [13]   // TEMPERATURE BREAKPOINT G. TIME 1/10 HOURS(ALWAYS=0)
        [3]   // TEMPERATURE BREAKPOINT B. TIME 1/10 HOURS(ALWAYS=0)
        [30].5   // Current vessel deferred chilling temp.high flag
        [30].3   // Current vessel deferred chilling active
        [5]   // TEMPERATURE BREAKPOINT C. TIME 1/10 HOURS(ALWAYS=0)
        [7]   // TEMPERATURE BREAKPOINT D. TIME 1/10 HOURS(ALWAYS=0)
        [9]   // TEMPERATURE BREAKPOINT E. TIME 1/10 HOURS(ALWAYS=0)
        [16].1   // Profile control flag Hold at B.P B
        [16].2   // Profile control flag Hold at B.P C
        [16].3   // Profile control flag Hold at B.P D
        [16].4   // Profile control flag Hold at B.P E
        [16].5   // Profile control flag Hold at B.P F
        [16].6   // Profile control flag Hold at B.P G
        [15].2   // PLC TO FOLLOW RAMP Breakpoints A to B
        [0]   // FV SYSTEM WORKING BUFFER VESSEL NUMBER
        [10]   // TEMPERATURE SETPOINT E. 1/10 DEGREE 'C'
        [12]   // TEMPERATURE SETPOINT F. 1/10 DEGREE 'C'
        [14]   // TEMPERATURE SETPOINT G. 1/10 DEGREE 'C'
        [21]   // Current vessel cold conditioning time
        [2]   // TEMPERATURE SETPOINT A. 1/10 DEGREE 'C'
        [30].4   // Current vessel final temp.reached
        [36]   // Current vessel time to deferred chlling start (hrs.x10)
        [4]   // TEMPERATURE SETPOINT B. 1/10 DEGREE 'C'
        [30].6   // Current vessel cold cond.temp.reached
        [6]   // TEMPERATURE SETPOINT C. 1/10 DEGREE 'C'
        [8]   // TEMPERATURE SETPOINT D. 1/10 DEGREE 'C'
        [15].3   // PLC TO USE CONE COOLING JACKET
        [25]   // ACTUAL TEMPERATURE -DEGREES 'C'*10
        [26]   // Calculated Setpoint 1/10 degrees C
        [44]   // Current vessel powder amount
        [20]   // Current FV warm conditioning time
        [29]   // FLAGS - PLC CONTROL
        [15]   // FLAGS-PROFILE CONTROL
        [28]   // CURRENT VOLUME HL*10
        [30].1   // Rouser required
        [27]   // CURRENT ELAPSED HOURS *10
        [30].0   // Cooling Valve to open
        [15].7   // PC>PLC Rousing enabled
        [43]   // Current vessel powder type
   MV_N111 : INT[50] := ([0] := 29, [2] := 80, [3] := 1200, [4] := 80, [5] := 1730, [6] := 80, [7] := 5040, [8] := 80, [9] := 6720, [10] := 80, [11] := 8400, [12] := 80, [13] := 32767, [14] := 80, [15] := 148, [17] := -32767, [18] := -32767, [19] := 1680, [20] := 311, [22] := 1947, [23] := 1, [24] := 10, [25] := 80, [26] := 80, [27] := 311, [30] := 19, [32] := 2, [34] := 2, [36] := 170, [42] := 25900);   // MV 1, CURRENT FV DATA
        [24]   // MV 1,Phase 0=off 8=Wait yeast 9=Wait Fill 10=Maturation 11to16=Conditioning
        [11]   // MV 1,TEMPERATURE BREAKPOINT F. TIME 1/10 HOURS(ALWAYS=0)
        [13]   // MV 1,TEMPERATURE BREAKPOINT G. TIME 1/10 HOURS(ALWAYS=0)
        [30].5   // MV 1,Current vessel deferred chilling temp.high flag
        [1]   // MV 1,TEMPERATURE BREAKPOINT A. TIME 1/10 HOURS(ALWAYS=0)
        [29].1   // MV 1,Current vessel deferred chilling enabled flag
        [3]   // MV 1,TEMPERATURE BREAKPOINT B. TIME 1/10 HOURS(ALWAYS=0)
        [5]   // MV 1,TEMPERATURE BREAKPOINT C. TIME 1/10 HOURS(ALWAYS=0)
        [36]   // MV 1,Current vessel time to deferred chlling start (hrs.x10)
        [15].5   // MV 1,Profile Control Flags : This is a Conditioning Profile
        [40]   // MV 1,Vessel RoutingStatus 0=Clean,1=Filling,2= Beer,3=Packng1,4=Pac kng2,5=Packng3,6=Ven ting,7=Dirty,8=CIP
        [15].7   // MV 1,PC>PLC Rousing enabled
        [43]   // MV 1,Current vessel powder type
        [15].4   // MV 1,Profile Control Flags : This is a Maturation Profile
        [16].1   // MV 1,Profile control flag Hold at B.P B
        [16].2   // MV 1,Profile control flag Hold at B.P C
        [10]   // MV 1,TEMPERATURE SETPOINT E. 1/10 DEGREE 'C'
        [7]   // MV 1,TEMPERATURE BREAKPOINT D. TIME 1/10 HOURS(ALWAYS=0)
        [12]   // MV 1,TEMPERATURE SETPOINT F. 1/10 DEGREE 'C'
        [14]   // MV 1,TEMPERATURE SETPOINT G. 1/10 DEGREE 'C'
        [9]   // MV 1,TEMPERATURE BREAKPOINT E. TIME 1/10 HOURS(ALWAYS=0)
        [0]   // MV 1,FV SYSTEM WORKING BUFFER VESSEL NUMBER
        [21]   // MV 1,Current vessel cold conditioning time
        [16].3   // MV 1,Profile control flag Hold at B.P D
        [2]   // MV 1,TEMPERATURE SETPOINT A. 1/10 DEGREE 'C'
        [30].3   // MV 1,Current vessel deferred chilling active
        [16].4   // MV 1,Profile control flag Hold at B.P E
        [30].4   // MV 1,Current vessel final temp.reached
        [16].5   // MV 1,Profile control flag Hold at B.P F
        [4]   // MV 1,TEMPERATURE SETPOINT B. 1/10 DEGREE 'C'
        [15].2   // MV 1,PLC TO FOLLOW RAMP Breakpoints A to B
        [20]   // MV 1,Current FV warm conditioning time
        [15].3   // MV 1,PLC TO USE CONE COOLING JACKET
        [15].9   // MV 1,Current vessel deferred chilling manual override
        [30].6   // MV 1,Current vessel cold cond.temp.reached
        [25]   // MV 1,ACTUAL TEMPERATURE -DEGREES 'C'*10
        [29]   // MV 1,FLAGS - PLC CONTROL
        [6]   // MV 1,TEMPERATURE SETPOINT C. 1/10 DEGREE 'C'
        [16].6   // MV 1,Profile control flag Hold at B.P G
        [30].1   // MV 1,Rouser required
        [27]   // MV 1,CURRENT ELAPSED HOURS *10
        [22]   // MV 1,Current FV total residence time
        [29].0   // MV 1,PC TO SAVE TEMPERATURE DATA
        [30].0   // MV 1,Cooling Valve to open
        [8]   // MV 1,TEMPERATURE SETPOINT D. 1/10 DEGREE 'C'
        [26]   // MV 1,Calculated Setpoint 1/10 degrees C
        [44]   // MV 1,Current vessel powder amount
        [28]   // MV 1,CURRENT VOLUME HL*10
        [15]   // MV 1,FLAGS-PROFILE CONTROL
   MV_N112 : INT[50] := ([0] := 30, [2] := 80, [3] := 1200, [4] := 80, [5] := 2050, [6] := 80, [7] := 5040, [8] := 80, [9] := 6720, [10] := 80, [11] := 8400, [12] := 80, [13] := 32767, [14] := 80, [15] := 148, [17] := -32767, [18] := -32767, [19] := 1680, [20] := 8251, [22] := 9870, [23] := 3, [24] := 10, [25] := 82, [26] := 80, [27] := 3383, [29] := 2, [30] := 24, [32] := 2, [34] := 2);   // MV 2, CURRENT FV DATA
